HMI tags "VAT_DB_SDC_EMS_FLAGS"
   "SDC\DB_SDC_EMS_FLAGS\DB_SDC_EMS_FLAGS.EMS[8]" : Int AT %DB0.DBW0, 1 s   // EMSdriver present
   "SDC\DB_SDC_EMS_FLAGS\_EMS_Flags_HMI_Byte_00" : Int, internal
   "SDC\DB_SDC_EMS_FLAGS\_EMS_Flags_HMI_Byte_19" : Int, internal
   "DB_SDC_EMS_FLAGS_HMI_HMI[1].RET_VAL_SFC12" : Int = PLC DB_SDC_EMS_FLAGS_HMI.HMI[1].RET_VAL_SFC12 AT %DB3801.DBW34, 1 s   // RetVal SFC12
   "SDC\DB_SDC_EMS_FLAGS\DB_SDC_EMS_FLAGS.EMS[9]" : Int AT %DB0.DBW0, 1 s   // EMSdriver present
   "SDC\DB_SDC_EMS_FLAGS\DB_SDC_EMS_FLAGS.EMS[19]" : Int AT %DB0.DBW0, 1 s   // EMSdriver present
   "SDC\DB_SDC_EMS_FLAGS\DB_SDC_EMS_FLAGS.HMI[XX].EMS_Nr" : Int AT %DB0.DBW0, 1 s   // Sektionsnummer
   "SDC\DB_SDC_EMS_FLAGS\_EMS_Flags_HMI_Byte_04" : Int, internal
   "SDC\DB_SDC_EMS_FLAGS\DB_SDC_EMS_FLAGS.HMI[XX].PULT_Nr_EDIT" : Int AT %DB0.DBW0, 1 s   // Pult Nr Editieren Aktiv (HMI 1 = Master)
   "SDC\DB_SDC_EMS_FLAGS\DB_SDC_EMS_FLAGS.EMS[20]" : Int AT %DB0.DBW0, 1 s   // EMSdriver present
   "DB_SDC_EMS_FLAGS_HEADER.LAENGE_EMS_FLAGS" : Int = PLC DB_SDC_EMS_FLAGS.HEADER.LAENGE_EMS_FLAGS AT %DB3701.DBW8, 1 s   // Länge Eingänge pro EMS
   "SDC\DB_SDC_EMS_FLAGS\DB_SDC_EMS_FLAGS.EMS[6]" : Int AT %DB0.DBW0, 1 s   // EMSdriver present
   "SDC\DB_SDC_EMS_FLAGS\DB_SDC_EMS_FLAGS.EMS[12]" : Int AT %DB0.DBW0, 1 s   // EMSdriver present
   "SDC\DB_SDC_EMS_FLAGS\DB_SDC_EMS_FLAGS.EMS[1]" : Int AT %DB0.DBW0, 1 s   // EMSdriver present
   "SDC\DB_SDC_EMS_FLAGS\DB_SDC_EMS_FLAGS.EMS[3]" : Int AT %DB0.DBW0, 1 s   // EMSdriver present
   "SDC\DB_SDC_EMS_FLAGS\DB_SDC_EMS_FLAGS.HMI[XX].BILD_Nr" : Int AT %DB0.DBW0, 1 s   // Bild_Nr aktiv
   "SDC\DB_SDC_EMS_FLAGS\DB_SDC_EMS_FLAGS.HMI[XX].T_LOAD" : Bool AT %DB0.DBX0.3, 1 s   // Taster laden
   "DB_SDC_EMS_FLAGS_HMI_HEADER.START_HMI" : Int = PLC DB_SDC_EMS_FLAGS_HMI.HEADER.START_HMI AT %DB3801.DBW10, 1 s   // Startadresse HMI
   "SDC\DB_SDC_EMS_FLAGS\DB_SDC_EMS_FLAGS.EMS[10]" : Int AT %DB0.DBW0, 1 s   // EMSdriver present
   "SDC\DB_SDC_EMS_FLAGS\_EMS_Flags_HMI_Byte_18" : Int, internal
   "SDC\DB_SDC_EMS_FLAGS\DB_SDC_EMS_FLAGS.EMS[7]" : Int AT %DB0.DBW0, 1 s   // EMSdriver present
   "SDC\DB_SDC_EMS_FLAGS\DB_SDC_EMS_FLAGS.EMS[13]" : Int AT %DB0.DBW0, 1 s   // EMSdriver present
   "DB_SDC_EMS_FLAGS_HMI_HMI[1].MODE_SFC12" : Byte = PLC DB_SDC_EMS_FLAGS_HMI.HMI[1].MODE_SFC12 AT %DB3801.DBB36, 1 s   // Mode SFC12
   "SDC\DB_SDC_EMS_FLAGS\DB_SDC_EMS_FLAGS.HMI[XX].FR_EDIT" : Bool AT %DB0.DBX0.0, 1 s   // Freigabe Editieren
   "SDC\DB_SDC_EMS_FLAGS\_EMS_Flags_HMI_Byte_12" : Int, internal
   "SDC\DB_SDC_EMS_FLAGS\DB_SDC_EMS_FLAGS.EMS[18]" : Int AT %DB0.DBW0, 1 s   // EMSdriver present
   "DB_SDC_EMS_FLAGS_HEADER.DB_NR" : Int = PLC DB_SDC_EMS_FLAGS.HEADER.DB_NR AT %DB3701.DBW0, 1 s   // DB Nummer
   "SDC\DB_SDC_EMS_FLAGS\DB_SDC_EMS_FLAGS.HMI[XX].BILD_Nr_Alt" : Int AT %DB0.DBW0, 1 s   // Bild_Nr alt
   "DB_SDC_EMS_FLAGS_HMI_HEADER.OFFEST_HMI_DATA" : Int = PLC DB_SDC_EMS_FLAGS_HMI.HEADER.OFFEST_HMI_DATA AT %DB3801.DBW12, 1 s   // Offestadresse der HMI Flag Data
   "SDC\DB_SDC_EMS_FLAGS\DB_SDC_EMS_FLAGS.EMS[2]" : Int AT %DB0.DBW0, 1 s   // EMSdriver present
   "DB_SDC_EMS_FLAGS_HEADER.MIN_NR_EMS" : Int = PLC DB_SDC_EMS_FLAGS.HEADER.MIN_NR_EMS AT %DB3701.DBW2, 1 s   // Niedrigste EMS Nummer im Daten DB
   "SDC\DB_SDC_EMS_FLAGS\DB_SDC_EMS_FLAGS.HMI[XX].T_ACTIV" : Bool AT %DB0.DBX0.4, 1 s   // Taster activieren
   "SDC\DB_SDC_EMS_FLAGS\DB_SDC_EMS_FLAGS.EMS[16]" : Int AT %DB0.DBW0, 1 s   // EMSdriver present
   "SDC\DB_SDC_EMS_FLAGS\DB_SDC_EMS_FLAGS.HMI[XX].T_DEACTIV" : Bool AT %DB0.DBX0.5, 1 s   // Taster deactivieren
   "DB_SDC_EMS_FLAGS_HEADER.MAX_NR_EMS" : Int = PLC DB_SDC_EMS_FLAGS.HEADER.MAX_NR_EMS AT %DB3701.DBW4, 1 s   // Höchste EMS Nummer im Daten DB
   "DB_SDC_EMS_FLAGS_HMI_HMI[1].REQ_SFC12" : Bool = PLC DB_SDC_EMS_FLAGS_HMI.HMI[1].REQ_SFC12 AT %DB3801.DBX39.3, 1 s   // Request SFC12
   "SDC\DB_SDC_EMS_FLAGS\DB_SDC_EMS_FLAGS.HMI[XX].T_RESET_BED" : Bool AT %DB0.DBX0.1, 1 s   // Taster Reset Bedienfreigabe Pult Nr Bedienung
   "SDC\DB_SDC_EMS_FLAGS\_EMS_Flags_HMI_Byte_20" : Int, internal
   "DB_SDC_EMS_FLAGS_HMI_HMI[1].PULT_Nr_EDIT" : Int = PLC DB_SDC_EMS_FLAGS_HMI.HMI[1].PULT_Nr_EDIT AT %DB3801.DBW20, 1 s   // Pult Nr Editieren Aktiv (HMI 1 = Master)
   "SDC\DB_SDC_EMS_FLAGS\DB_SDC_EMS_FLAGS.HMI[XX].ER_DATA" : Bool AT %DB0.DBX0.1, 1 s   // Daten Fehlerhaft
   "SDC\DB_SDC_EMS_FLAGS\_EMS_Flags_HMI_Byte_08" : Int, internal
   "SDC\DB_SDC_EMS_FLAGS\DB_SDC_EMS_FLAGS.EMS[11]" : Int AT %DB0.DBW0, 1 s   // EMSdriver present
   "DB_SDC_EMS_FLAGS_HMI_HMI[1].TIME_SFC12" : Int = PLC DB_SDC_EMS_FLAGS_HMI.HMI[1].TIME_SFC12 AT %DB3801.DBW30, 1 s   // Actuelle Zeit Activieren/Deactivieren
   "SDC\DB_SDC_EMS_FLAGS\DB_SDC_EMS_FLAGS.EMS[14]" : Int AT %DB0.DBW0, 1 s   // EMSdriver present
   "SDC\DB_SDC_EMS_FLAGS\_EMS_Flags_HMI_Byte_16" : Int, internal
   "SDC\DB_SDC_EMS_FLAGS\DB_SDC_EMS_FLAGS.HMI[XX].T_SAVE" : Bool AT %DB0.DBX0.2, 1 s   // Taster speichern
   "SDC\DB_SDC_EMS_FLAGS\DB_SDC_EMS_FLAGS.EMS[15]" : Int AT %DB0.DBW0, 1 s   // EMSdriver present
   "SDC\DB_SDC_EMS_FLAGS\_EMS_Flags_HMI_Byte_10" : Int, internal
   "SDC\DB_SDC_EMS_FLAGS\_EMS_Flags_HMI_Byte_14" : Int, internal
   "SDC\DB_SDC_EMS_FLAGS\DB_SDC_EMS_FLAGS.HMI[XX].T_EDIT" : Bool AT %DB0.DBX0.0, 1 s   // Taster Editieren für Pult aktivieren
   "SDC\DB_SDC_EMS_FLAGS\_EMS_Flags_HMI_Byte_09" : Int, internal
   "DB_SDC_EMS_FLAGS_HMI_HMI[1].BUSY_SFC12" : Bool = PLC DB_SDC_EMS_FLAGS_HMI.HMI[1].BUSY_SFC12 AT %DB3801.DBX39.2, 1 s   // Busy SFC12
   "SDC\DB_SDC_EMS_FLAGS\_EMS_Nr" : Int, internal
      on ChangeValue: "SDC_TS_PARAMETER"(); "SDC_TS_REFERENCE"("SDC\DB_SDC_EMS_FLAGS\_EMS_Nr")
   "SDC\DB_SDC_EMS_FLAGS\DB_SDC_EMS_FLAGS.EMS[17]" : Int AT %DB0.DBW0, 1 s   // EMSdriver present
   "SDC\DB_SDC_EMS_FLAGS\_EMS_Flags_HMI_Byte_06" : Int, internal
   "SDC\DB_SDC_EMS_FLAGS\DB_SDC_EMS_FLAGS.HMI[XX].FLAGS" : Word AT %DB0.DBW0, 1 s   // Freigabe Editieren
   "SDC\DB_SDC_EMS_FLAGS\_EMS_Flags_HMI_Byte_02" : Int, internal
   "SDC\DB_SDC_EMS_FLAGS\DB_SDC_EMS_FLAGS.EMS[5]" : Int AT %DB0.DBW0, 1 s   // EMSdriver present
   "DB_SDC_EMS_FLAGS_HEADER.START_EMS" : Int = PLC DB_SDC_EMS_FLAGS.HEADER.START_EMS AT %DB3701.DBW6, 1 s   // Startadresse der EMS Daten im Daten DB
   "SDC\DB_SDC_EMS_FLAGS\DB_SDC_EMS_FLAGS.EMS[4]" : Int AT %DB0.DBW0, 1 s   // EMSdriver present
   "SDC\DB_SDC_EMS_FLAGS\DB_SDC_EMS_FLAGS.HMI[1].LADDR_SFC12" : Int AT %DB0.DBW32, 1 s   // Actuelle LADDR
   "SDC\DB_SDC_EMS_FLAGS\DB_SDC_EMS_FLAGS.EMS[21]" : Int AT %DB0.DBW0, 1 s   // EMSdriver present
   "SDC\DB_SDC_EMS_FLAGS\DB_SDC_EMS_FLAGS.EMS[22]" : Int AT %DB0.DBW0, 1 s
   "SDC\DB_SDC_EMS_FLAGS\DB_SDC_EMS_FLAGS.EMS[23]" : Int AT %DB0.DBW0, 1 s
   "SDC\DB_SDC_EMS_FLAGS\DB_SDC_EMS_FLAGS.EMS[24]" : Int AT %DB0.DBW0, 1 s
   "SDC\DB_SDC_EMS_FLAGS\DB_SDC_EMS_FLAGS.EMS[25]" : Int AT %DB0.DBW0, 1 s
   "SDC\DB_SDC_EMS_FLAGS\DB_SDC_EMS_FLAGS.EMS[26]" : Int AT %DB0.DBW0, 1 s
   "SDC\DB_SDC_EMS_FLAGS\DB_SDC_EMS_FLAGS.EMS[27]" : Int AT %DB0.DBW0, 1 s
   "SDC\DB_SDC_EMS_FLAGS\DB_SDC_EMS_FLAGS.EMS[28]" : Int AT %DB0.DBW0, 1 s
   "SDC\DB_SDC_EMS_FLAGS\DB_SDC_EMS_FLAGS.EMS[29]" : Int AT %DB0.DBW0, 1 s
   "SDC\DB_SDC_EMS_FLAGS\DB_SDC_EMS_FLAGS.EMS[30]" : Int AT %DB0.DBW0, 1 s
   "SDC\DB_SDC_EMS_FLAGS\DB_SDC_EMS_FLAGS.EMS[31]" : Int AT %DB0.DBW0, 1 s
   "SDC\DB_SDC_EMS_FLAGS\DB_SDC_EMS_FLAGS.EMS[32]" : Int AT %DB0.DBW0, 1 s
   "SDC\DB_SDC_EMS_FLAGS\DB_SDC_EMS_FLAGS.EMS[33]" : Int AT %DB0.DBW0, 1 s
   "SDC\DB_SDC_EMS_FLAGS\DB_SDC_EMS_FLAGS.EMS[34]" : Int AT %DB0.DBW0, 1 s
   "SDC\DB_SDC_EMS_FLAGS\DB_SDC_EMS_FLAGS.EMS[35]" : Int AT %DB0.DBW0, 1 s
   "SDC\DB_SDC_EMS_FLAGS\DB_SDC_EMS_FLAGS.EMS[36]" : Int AT %DB0.DBW0, 1 s
   "SDC\DB_SDC_EMS_FLAGS\DB_SDC_EMS_FLAGS.EMS[37]" : Int AT %DB0.DBW0, 1 s
   "SDC\DB_SDC_EMS_FLAGS\DB_SDC_EMS_FLAGS.EMS[38]" : Int AT %DB0.DBW0, 1 s
   "SDC\DB_SDC_EMS_FLAGS\DB_SDC_EMS_FLAGS.EMS[39]" : Int AT %DB0.DBW0, 1 s
   "SDC\DB_SDC_EMS_FLAGS\DB_SDC_EMS_FLAGS.EMS[40]" : Int AT %DB0.DBW0, 1 s
   "SDC\DB_SDC_EMS_FLAGS\DB_SDC_EMS_FLAGS.EMS[41]" : Int AT %DB0.DBW0, 1 s
   "SDC\DB_SDC_EMS_FLAGS\DB_SDC_EMS_FLAGS.EMS[42]" : Int AT %DB0.DBW0, 1 s
   "SDC\DB_SDC_EMS_FLAGS\DB_SDC_EMS_FLAGS.EMS[43]" : Int AT %DB0.DBW0, 1 s
   "SDC\DB_SDC_EMS_FLAGS\DB_SDC_EMS_FLAGS.EMS[44]" : Int AT %DB0.DBW0, 1 s
   "SDC\DB_SDC_EMS_FLAGS\DB_SDC_EMS_FLAGS.EMS[45]" : Int AT %DB0.DBW0, 1 s
   "SDC\DB_SDC_EMS_FLAGS\DB_SDC_EMS_FLAGS.EMS[46]" : Int AT %DB0.DBW0, 1 s
   "SDC\DB_SDC_EMS_FLAGS\DB_SDC_EMS_FLAGS.EMS[47]" : Int AT %DB0.DBW0, 1 s
   "SDC\DB_SDC_EMS_FLAGS\DB_SDC_EMS_FLAGS.EMS[48]" : Int AT %DB0.DBW0, 1 s
   "SDC\DB_SDC_EMS_FLAGS\DB_SDC_EMS_FLAGS.EMS[49]" : Int AT %DB0.DBW0, 1 s
   "SDC\DB_SDC_EMS_FLAGS\DB_SDC_EMS_FLAGS.EMS[50]" : Int AT %DB0.DBW0, 1 s
   "SDC\DB_SDC_EMS_FLAGS\DB_SDC_EMS_FLAGS.EMS[51]" : Int AT %DB0.DBW0, 1 s
   "SDC\DB_SDC_EMS_FLAGS\DB_SDC_EMS_FLAGS.EMS[52]" : Int AT %DB0.DBW0, 1 s
   "SDC\DB_SDC_EMS_FLAGS\DB_SDC_EMS_FLAGS.EMS[53]" : Int AT %DB0.DBW0, 1 s
   "SDC\DB_SDC_EMS_FLAGS\DB_SDC_EMS_FLAGS.EMS[54]" : Int AT %DB0.DBW0, 1 s
   "SDC\DB_SDC_EMS_FLAGS\DB_SDC_EMS_FLAGS.EMS[55]" : Int AT %DB0.DBW0, 1 s
   "SDC\DB_SDC_EMS_FLAGS\DB_SDC_EMS_FLAGS.EMS[56]" : Int AT %DB0.DBW0, 1 s
   "SDC\DB_SDC_EMS_FLAGS\DB_SDC_EMS_FLAGS.EMS[57]" : Int AT %DB0.DBW0, 1 s
   "SDC\DB_SDC_EMS_FLAGS\DB_SDC_EMS_FLAGS.EMS[58]" : Int AT %DB0.DBW0, 1 s
   "SDC\DB_SDC_EMS_FLAGS\DB_SDC_EMS_FLAGS.EMS[59]" : Int AT %DB0.DBW0, 1 s
   "SDC\DB_SDC_EMS_FLAGS\DB_SDC_EMS_FLAGS.EMS[60]" : Int AT %DB0.DBW0, 1 s
   "SDC\DB_SDC_EMS_FLAGS\DB_SDC_EMS_FLAGS.EMS[61]" : Int AT %DB0.DBW0, 1 s
   "SDC\DB_SDC_EMS_FLAGS\DB_SDC_EMS_FLAGS.EMS[62]" : Int AT %DB0.DBW0, 1 s
   "SDC\DB_SDC_EMS_FLAGS\DB_SDC_EMS_FLAGS.EMS[63]" : Int AT %DB0.DBW0, 1 s
   "SDC\DB_SDC_EMS_FLAGS\DB_SDC_EMS_FLAGS.EMS[64]" : Int AT %DB0.DBW0, 1 s
   "SDC\DB_SDC_EMS_FLAGS\DB_SDC_EMS_FLAGS.EMS[65]" : Int AT %DB0.DBW0, 1 s
   "SDC\DB_SDC_EMS_FLAGS\DB_SDC_EMS_FLAGS.EMS[66]" : Int AT %DB0.DBW0, 1 s
   "SDC\DB_SDC_EMS_FLAGS\DB_SDC_EMS_FLAGS.EMS[67]" : Int AT %DB0.DBW0, 1 s
   "SDC\DB_SDC_EMS_FLAGS\DB_SDC_EMS_FLAGS.EMS[68]" : Int AT %DB0.DBW0, 1 s
   "SDC\DB_SDC_EMS_FLAGS\DB_SDC_EMS_FLAGS.EMS[69]" : Int AT %DB0.DBW0, 1 s
   "SDC\DB_SDC_EMS_FLAGS\DB_SDC_EMS_FLAGS.EMS[70]" : Int AT %DB0.DBW0, 1 s
   "SDC\DB_SDC_EMS_FLAGS\DB_SDC_EMS_FLAGS.EMS[71]" : Int AT %DB0.DBW0, 1 s
   "SDC\DB_SDC_EMS_FLAGS\DB_SDC_EMS_FLAGS.EMS[72]" : Int AT %DB0.DBW0, 1 s
   "SDC\DB_SDC_EMS_FLAGS\DB_SDC_EMS_FLAGS.EMS[73]" : Int AT %DB0.DBW0, 1 s
   "SDC\DB_SDC_EMS_FLAGS\DB_SDC_EMS_FLAGS.EMS[74]" : Int AT %DB0.DBW0, 1 s
   "SDC\DB_SDC_EMS_FLAGS\DB_SDC_EMS_FLAGS.EMS[75]" : Int AT %DB0.DBW0, 1 s
   "SDC\DB_SDC_EMS_FLAGS\DB_SDC_EMS_FLAGS.EMS[76]" : Int AT %DB0.DBW0, 1 s
   "SDC\DB_SDC_EMS_FLAGS\DB_SDC_EMS_FLAGS.EMS[77]" : Int AT %DB0.DBW0, 1 s
   "SDC\DB_SDC_EMS_FLAGS\DB_SDC_EMS_FLAGS.EMS[78]" : Int AT %DB0.DBW0, 1 s
   "SDC\DB_SDC_EMS_FLAGS\DB_SDC_EMS_FLAGS.EMS[79]" : Int AT %DB0.DBW0, 1 s
   "SDC\DB_SDC_EMS_FLAGS\DB_SDC_EMS_FLAGS.EMS[80]" : Int AT %DB0.DBW0, 1 s
   "SDC\DB_SDC_EMS_FLAGS\DB_SDC_EMS_FLAGS.EMS[81]" : Int AT %DB0.DBW0, 1 s
   "SDC\DB_SDC_EMS_FLAGS\DB_SDC_EMS_FLAGS.EMS[82]" : Int AT %DB0.DBW0, 1 s
   "SDC\DB_SDC_EMS_FLAGS\DB_SDC_EMS_FLAGS.EMS[83]" : Int AT %DB0.DBW0, 1 s
   "SDC\DB_SDC_EMS_FLAGS\DB_SDC_EMS_FLAGS.EMS[84]" : Int AT %DB0.DBW0, 1 s
   "SDC\DB_SDC_EMS_FLAGS\DB_SDC_EMS_FLAGS.EMS[85]" : Int AT %DB0.DBW0, 1 s
   "SDC\DB_SDC_EMS_FLAGS\DB_SDC_EMS_FLAGS.EMS[86]" : Int AT %DB0.DBW0, 1 s
   "SDC\DB_SDC_EMS_FLAGS\DB_SDC_EMS_FLAGS.EMS[87]" : Int AT %DB0.DBW0, 1 s
   "SDC\DB_SDC_EMS_FLAGS\DB_SDC_EMS_FLAGS.EMS[88]" : Int AT %DB0.DBW0, 1 s
   "SDC\DB_SDC_EMS_FLAGS\DB_SDC_EMS_FLAGS.EMS[89]" : Int AT %DB0.DBW0, 1 s
   "SDC\DB_SDC_EMS_FLAGS\DB_SDC_EMS_FLAGS.EMS[90]" : Int AT %DB0.DBW0, 1 s
   "SDC\DB_SDC_EMS_FLAGS\DB_SDC_EMS_FLAGS.EMS[91]" : Int AT %DB0.DBW0, 1 s
   "SDC\DB_SDC_EMS_FLAGS\DB_SDC_EMS_FLAGS.EMS[92]" : Int AT %DB0.DBW0, 1 s
   "SDC\DB_SDC_EMS_FLAGS\DB_SDC_EMS_FLAGS.EMS[93]" : Int AT %DB0.DBW0, 1 s
   "SDC\DB_SDC_EMS_FLAGS\DB_SDC_EMS_FLAGS.EMS[94]" : Int AT %DB0.DBW0, 1 s
   "SDC\DB_SDC_EMS_FLAGS\DB_SDC_EMS_FLAGS.EMS[95]" : Int AT %DB0.DBW0, 1 s
   "SDC\DB_SDC_EMS_FLAGS\DB_SDC_EMS_FLAGS.EMS[96]" : Int AT %DB0.DBW0, 1 s
   "SDC\DB_SDC_EMS_FLAGS\DB_SDC_EMS_FLAGS.EMS[97]" : Int AT %DB0.DBW0, 1 s
   "SDC\DB_SDC_EMS_FLAGS\DB_SDC_EMS_FLAGS.EMS[98]" : Int AT %DB0.DBW0, 1 s
   "SDC\DB_SDC_EMS_FLAGS\DB_SDC_EMS_FLAGS.EMS[99]" : Int AT %DB0.DBW0, 1 s
   "SDC\DB_SDC_EMS_FLAGS\DB_SDC_EMS_FLAGS.EMS[100]" : Int AT %DB0.DBW0, 1 s
   "SDC\DB_SDC_EMS_FLAGS\DB_SDC_EMS_FLAGS.EMS[101]" : Int AT %DB0.DBW0, 1 s
   "SDC\DB_SDC_EMS_FLAGS\DB_SDC_EMS_FLAGS.EMS[102]" : Int AT %DB0.DBW0, 1 s
   "SDC\DB_SDC_EMS_FLAGS\DB_SDC_EMS_FLAGS.EMS[103]" : Int AT %DB0.DBW0, 1 s
   "SDC\DB_SDC_EMS_FLAGS\DB_SDC_EMS_FLAGS.EMS[104]" : Int AT %DB0.DBW0, 1 s
   "SDC\DB_SDC_EMS_FLAGS\DB_SDC_EMS_FLAGS.EMS[105]" : Int AT %DB0.DBW0, 1 s
   "SDC\DB_SDC_EMS_FLAGS\DB_SDC_EMS_FLAGS.EMS[106]" : Int AT %DB0.DBW0, 1 s
   "SDC\DB_SDC_EMS_FLAGS\DB_SDC_EMS_FLAGS.EMS[107]" : Int AT %DB0.DBW0, 1 s
   "SDC\DB_SDC_EMS_FLAGS\DB_SDC_EMS_FLAGS.EMS[108]" : Int AT %DB0.DBW0, 1 s
   "SDC\DB_SDC_EMS_FLAGS\DB_SDC_EMS_FLAGS.EMS[109]" : Int AT %DB0.DBW0, 1 s
   "SDC\DB_SDC_EMS_FLAGS\_EMS_Flags_Byte_EMS001" : Int, internal
   "SDC\DB_SDC_EMS_FLAGS\_EMS_Flags_Byte_EMS002" : Int, internal
   "SDC\DB_SDC_EMS_FLAGS\_EMS_Flags_Byte_EMS003" : Int, internal
   "SDC\DB_SDC_EMS_FLAGS\_EMS_Flags_Byte_EMS004" : Int, internal
   "SDC\DB_SDC_EMS_FLAGS\_EMS_Flags_Byte_EMS005" : Int, internal
   "SDC\DB_SDC_EMS_FLAGS\_EMS_Flags_Byte_EMS006" : Int, internal
   "SDC\DB_SDC_EMS_FLAGS\_EMS_Flags_Byte_EMS007" : Int, internal
   "SDC\DB_SDC_EMS_FLAGS\_EMS_Flags_Byte_EMS008" : Int, internal
   "SDC\DB_SDC_EMS_FLAGS\_EMS_Flags_Byte_EMS009" : Int, internal
   "SDC\DB_SDC_EMS_FLAGS\_EMS_Flags_Byte_EMS010" : Int, internal
   "SDC\DB_SDC_EMS_FLAGS\_EMS_Flags_Byte_EMS011" : Int, internal
   "SDC\DB_SDC_EMS_FLAGS\_EMS_Flags_Byte_EMS012" : Int, internal
   "SDC\DB_SDC_EMS_FLAGS\_EMS_Flags_Byte_EMS013" : Int, internal
   "SDC\DB_SDC_EMS_FLAGS\_EMS_Flags_Byte_EMS014" : Int, internal
   "SDC\DB_SDC_EMS_FLAGS\_EMS_Flags_Byte_EMS015" : Int, internal
   "SDC\DB_SDC_EMS_FLAGS\_EMS_Flags_Byte_EMS016" : Int, internal
   "SDC\DB_SDC_EMS_FLAGS\_EMS_Flags_Byte_EMS017" : Int, internal
   "SDC\DB_SDC_EMS_FLAGS\_EMS_Flags_Byte_EMS018" : Int, internal
   "SDC\DB_SDC_EMS_FLAGS\_EMS_Flags_Byte_EMS019" : Int, internal
   "SDC\DB_SDC_EMS_FLAGS\_EMS_Flags_Byte_EMS020" : Int, internal
   "SDC\DB_SDC_EMS_FLAGS\_EMS_Flags_Byte_EMS021" : Int, internal
   "SDC\DB_SDC_EMS_FLAGS\_EMS_Flags_Byte_EMS022" : Int, internal
   "SDC\DB_SDC_EMS_FLAGS\_EMS_Flags_Byte_EMS023" : Int, internal
   "SDC\DB_SDC_EMS_FLAGS\_EMS_Flags_Byte_EMS024" : Int, internal
   "SDC\DB_SDC_EMS_FLAGS\_EMS_Flags_Byte_EMS025" : Int, internal
   "SDC\DB_SDC_EMS_FLAGS\_EMS_Flags_Byte_EMS026" : Int, internal
   "SDC\DB_SDC_EMS_FLAGS\_EMS_Flags_Byte_EMS027" : Int, internal
   "SDC\DB_SDC_EMS_FLAGS\_EMS_Flags_Byte_EMS028" : Int, internal
   "SDC\DB_SDC_EMS_FLAGS\_EMS_Flags_Byte_EMS029" : Int, internal
   "SDC\DB_SDC_EMS_FLAGS\_EMS_Flags_Byte_EMS030" : Int, internal
   "SDC\DB_SDC_EMS_FLAGS\_EMS_Flags_Byte_EMS031" : Int, internal
   "SDC\DB_SDC_EMS_FLAGS\_EMS_Flags_Byte_EMS032" : Int, internal
   "SDC\DB_SDC_EMS_FLAGS\_EMS_Flags_Byte_EMS033" : Int, internal
   "SDC\DB_SDC_EMS_FLAGS\_EMS_Flags_Byte_EMS034" : Int, internal
   "SDC\DB_SDC_EMS_FLAGS\_EMS_Flags_Byte_EMS035" : Int, internal
   "SDC\DB_SDC_EMS_FLAGS\_EMS_Flags_Byte_EMS036" : Int, internal
   "SDC\DB_SDC_EMS_FLAGS\_EMS_Flags_Byte_EMS037" : Int, internal
   "SDC\DB_SDC_EMS_FLAGS\_EMS_Flags_Byte_EMS038" : Int, internal
   "SDC\DB_SDC_EMS_FLAGS\_EMS_Flags_Byte_EMS039" : Int, internal
   "SDC\DB_SDC_EMS_FLAGS\_EMS_Flags_Byte_EMS040" : Int, internal
   "SDC\DB_SDC_EMS_FLAGS\_EMS_Flags_Byte_EMS041" : Int, internal
   "SDC\DB_SDC_EMS_FLAGS\_EMS_Flags_Byte_EMS042" : Int, internal
   "SDC\DB_SDC_EMS_FLAGS\_EMS_Flags_Byte_EMS043" : Int, internal
   "SDC\DB_SDC_EMS_FLAGS\_EMS_Flags_Byte_EMS044" : Int, internal
   "SDC\DB_SDC_EMS_FLAGS\_EMS_Flags_Byte_EMS045" : Int, internal
   "SDC\DB_SDC_EMS_FLAGS\_EMS_Flags_Byte_EMS046" : Int, internal
   "SDC\DB_SDC_EMS_FLAGS\_EMS_Flags_Byte_EMS047" : Int, internal
   "SDC\DB_SDC_EMS_FLAGS\_EMS_Flags_Byte_EMS048" : Int, internal
   "SDC\DB_SDC_EMS_FLAGS\_EMS_Flags_Byte_EMS049" : Int, internal
   "SDC\DB_SDC_EMS_FLAGS\_EMS_Flags_Byte_EMS050" : Int, internal
   "SDC\DB_SDC_EMS_FLAGS\_EMS_Flags_Byte_EMS051" : Int, internal
   "SDC\DB_SDC_EMS_FLAGS\_EMS_Flags_Byte_EMS052" : Int, internal
   "SDC\DB_SDC_EMS_FLAGS\_EMS_Flags_Byte_EMS053" : Int, internal
   "SDC\DB_SDC_EMS_FLAGS\_EMS_Flags_Byte_EMS054" : Int, internal
   "SDC\DB_SDC_EMS_FLAGS\_EMS_Flags_Byte_EMS055" : Int, internal
   "SDC\DB_SDC_EMS_FLAGS\_EMS_Flags_Byte_EMS056" : Int, internal
   "SDC\DB_SDC_EMS_FLAGS\_EMS_Flags_Byte_EMS057" : Int, internal
   "SDC\DB_SDC_EMS_FLAGS\_EMS_Flags_Byte_EMS058" : Int, internal
   "SDC\DB_SDC_EMS_FLAGS\_EMS_Flags_Byte_EMS059" : Int, internal
   "SDC\DB_SDC_EMS_FLAGS\_EMS_Flags_Byte_EMS060" : Int, internal
   "SDC\DB_SDC_EMS_FLAGS\_EMS_Flags_Byte_EMS061" : Int, internal
   "SDC\DB_SDC_EMS_FLAGS\_EMS_Flags_Byte_EMS062" : Int, internal
   "SDC\DB_SDC_EMS_FLAGS\_EMS_Flags_Byte_EMS063" : Int, internal
   "SDC\DB_SDC_EMS_FLAGS\_EMS_Flags_Byte_EMS064" : Int, internal
   "SDC\DB_SDC_EMS_FLAGS\_EMS_Flags_Byte_EMS065" : Int, internal
   "SDC\DB_SDC_EMS_FLAGS\_EMS_Flags_Byte_EMS066" : Int, internal
   "SDC\DB_SDC_EMS_FLAGS\_EMS_Flags_Byte_EMS067" : Int, internal
   "SDC\DB_SDC_EMS_FLAGS\_EMS_Flags_Byte_EMS068" : Int, internal
   "SDC\DB_SDC_EMS_FLAGS\_EMS_Flags_Byte_EMS069" : Int, internal
   "SDC\DB_SDC_EMS_FLAGS\_EMS_Flags_Byte_EMS070" : Int, internal
   "SDC\DB_SDC_EMS_FLAGS\_EMS_Flags_Byte_EMS071" : Int, internal
   "SDC\DB_SDC_EMS_FLAGS\_EMS_Flags_Byte_EMS072" : Int, internal
   "SDC\DB_SDC_EMS_FLAGS\_EMS_Flags_Byte_EMS073" : Int, internal
   "SDC\DB_SDC_EMS_FLAGS\_EMS_Flags_Byte_EMS074" : Int, internal
   "SDC\DB_SDC_EMS_FLAGS\_EMS_Flags_Byte_EMS075" : Int, internal
   "SDC\DB_SDC_EMS_FLAGS\_EMS_Flags_Byte_EMS076" : Int, internal
   "SDC\DB_SDC_EMS_FLAGS\_EMS_Flags_Byte_EMS077" : Int, internal
   "SDC\DB_SDC_EMS_FLAGS\_EMS_Flags_Byte_EMS078" : Int, internal
   "SDC\DB_SDC_EMS_FLAGS\_EMS_Flags_Byte_EMS079" : Int, internal
   "SDC\DB_SDC_EMS_FLAGS\_EMS_Flags_Byte_EMS080" : Int, internal
   "SDC\DB_SDC_EMS_FLAGS\_EMS_Flags_Byte_EMS081" : Int, internal
   "SDC\DB_SDC_EMS_FLAGS\_EMS_Flags_Byte_EMS082" : Int, internal
   "SDC\DB_SDC_EMS_FLAGS\_EMS_Flags_Byte_EMS083" : Int, internal
   "SDC\DB_SDC_EMS_FLAGS\_EMS_Flags_Byte_EMS084" : Int, internal
   "SDC\DB_SDC_EMS_FLAGS\_EMS_Flags_Byte_EMS085" : Int, internal
   "SDC\DB_SDC_EMS_FLAGS\_EMS_Flags_Byte_EMS086" : Int, internal
   "SDC\DB_SDC_EMS_FLAGS\_EMS_Flags_Byte_EMS087" : Int, internal
   "SDC\DB_SDC_EMS_FLAGS\_EMS_Flags_Byte_EMS088" : Int, internal
   "SDC\DB_SDC_EMS_FLAGS\_EMS_Flags_Byte_EMS089" : Int, internal
   "SDC\DB_SDC_EMS_FLAGS\_EMS_Flags_Byte_EMS090" : Int, internal
   "SDC\DB_SDC_EMS_FLAGS\_EMS_Flags_Byte_EMS091" : Int, internal
   "SDC\DB_SDC_EMS_FLAGS\_EMS_Flags_Byte_EMS092" : Int, internal
   "SDC\DB_SDC_EMS_FLAGS\_EMS_Flags_Byte_EMS093" : Int, internal
   "SDC\DB_SDC_EMS_FLAGS\_EMS_Flags_Byte_EMS094" : Int, internal
   "SDC\DB_SDC_EMS_FLAGS\_EMS_Flags_Byte_EMS095" : Int, internal
   "SDC\DB_SDC_EMS_FLAGS\_EMS_Flags_Byte_EMS096" : Int, internal
   "SDC\DB_SDC_EMS_FLAGS\_EMS_Flags_Byte_EMS097" : Int, internal
   "SDC\DB_SDC_EMS_FLAGS\_EMS_Flags_Byte_EMS098" : Int, internal
   "SDC\DB_SDC_EMS_FLAGS\_EMS_Flags_Byte_EMS099" : Int, internal
   "SDC\DB_SDC_EMS_FLAGS\_EMS_Flags_Byte_EMS100" : Int, internal
   "SDC\DB_SDC_EMS_FLAGS\_EMS_Flags_Byte_EMS101" : Int, internal
   "SDC\DB_SDC_EMS_FLAGS\_EMS_Flags_Byte_EMS102" : Int, internal
   "SDC\DB_SDC_EMS_FLAGS\_EMS_Flags_Byte_EMS103" : Int, internal
   "SDC\DB_SDC_EMS_FLAGS\_EMS_Flags_Byte_EMS104" : Int, internal
   "SDC\DB_SDC_EMS_FLAGS\_EMS_Flags_Byte_EMS105" : Int, internal
   "SDC\DB_SDC_EMS_FLAGS\_EMS_Flags_Byte_EMS106" : Int, internal
   "SDC\DB_SDC_EMS_FLAGS\_EMS_Flags_Byte_EMS107" : Int, internal
   "SDC\DB_SDC_EMS_FLAGS\_EMS_Flags_Byte_EMS108" : Int, internal
   "SDC\DB_SDC_EMS_FLAGS\_EMS_Flags_Byte_EMS109" : Int, internal
   "DB_SDC_EMS_FLAGS_HMI_HEADER.DB_NR" : Int = PLC DB_SDC_EMS_FLAGS_HMI.HEADER.DB_NR AT %DB3801.DBW0, 1 s
   "SDC\DB_SDC_EMS_FLAGS\_EMS_Flags_Byte_EMS110" : Int, internal
   "SDC\DB_SDC_EMS_FLAGS\_EMS_Flags_Byte_EMS111" : Int, internal
   "SDC\DB_SDC_EMS_FLAGS\_EMS_Flags_Byte_EMS112" : Int, internal
   "SDC\DB_SDC_EMS_FLAGS\_EMS_Flags_Byte_EMS113" : Int, internal
   "SDC\DB_SDC_EMS_FLAGS\_EMS_Flags_Byte_EMS114" : Int, internal
   "SDC\DB_SDC_EMS_FLAGS\_EMS_Flags_Byte_EMS115" : Int, internal
   "SDC\DB_SDC_EMS_FLAGS\_EMS_Flags_Byte_EMS116" : Int, internal
   "SDC\DB_SDC_EMS_FLAGS\_EMS_Flags_Byte_EMS117" : Int, internal
   "SDC\DB_SDC_EMS_FLAGS\_EMS_Flags_Byte_EMS118" : Int, internal
   "SDC\DB_SDC_EMS_FLAGS\_EMS_Flags_Byte_EMS119" : Int, internal
   "SDC\DB_SDC_EMS_FLAGS\_EMS_Flags_Byte_EMS120" : Int, internal
   "SDC\DB_SDC_EMS_FLAGS\_EMS_Flags_Byte_EMS121" : Int, internal
   "SDC\DB_SDC_EMS_FLAGS\_EMS_Flags_Byte_EMS122" : Int, internal
   "SDC\DB_SDC_EMS_FLAGS\_EMS_Flags_Byte_EMS123" : Int, internal
   "SDC\DB_SDC_EMS_FLAGS\_EMS_Flags_Byte_EMS124" : Int, internal
   "SDC\DB_SDC_EMS_FLAGS\_EMS_Flags_Byte_EMS125" : Int, internal
   "SDC\DB_SDC_EMS_FLAGS\_EMS_Flags_Byte_EMS126" : Int, internal
   "SDC\DB_SDC_EMS_FLAGS\_EMS_Flags_Byte_EMS127" : Int, internal
   "SDC\DB_SDC_EMS_FLAGS\_EMS_Flags_Byte_EMS128" : Int, internal
   "SDC\DB_SDC_EMS_FLAGS\_EMS_Flags_Byte_EMS129" : Int, internal
   "SDC\DB_SDC_EMS_FLAGS\_EMS_Flags_Byte_EMS130" : Int, internal
   "SDC\DB_SDC_EMS_FLAGS\_EMS_Flags_Byte_EMS131" : Int, internal
   "SDC\DB_SDC_EMS_FLAGS\_EMS_Flags_Byte_EMS132" : Int, internal
   "SDC\DB_SDC_EMS_FLAGS\_EMS_Flags_Byte_EMS133" : Int, internal
   "SDC\DB_SDC_EMS_FLAGS\_EMS_Flags_Byte_EMS134" : Int, internal
   "SDC\DB_SDC_EMS_FLAGS\_EMS_Flags_Byte_EMS135" : Int, internal
   "SDC\DB_SDC_EMS_FLAGS\_EMS_Flags_Byte_EMS136" : Int, internal
   "SDC\DB_SDC_EMS_FLAGS\_EMS_Flags_Byte_EMS137" : Int, internal
   "SDC\DB_SDC_EMS_FLAGS\_EMS_Flags_Byte_EMS138" : Int, internal
   "SDC\DB_SDC_EMS_FLAGS\_EMS_Flags_Byte_EMS139" : Int, internal
   "SDC\DB_SDC_EMS_FLAGS\_EMS_Flags_Byte_EMS140" : Int, internal
   "SDC\DB_SDC_EMS_FLAGS\_EMS_Flags_Byte_EMS141" : Int, internal
   "SDC\DB_SDC_EMS_FLAGS\_EMS_Flags_Byte_EMS142" : Int, internal
   "SDC\DB_SDC_EMS_FLAGS\_EMS_Flags_Byte_EMS143" : Int, internal
   "SDC\DB_SDC_EMS_FLAGS\_EMS_Flags_Byte_EMS144" : Int, internal
   "SDC\DB_SDC_EMS_FLAGS\_EMS_Flags_Byte_EMS145" : Int, internal
   "SDC\DB_SDC_EMS_FLAGS\_EMS_Flags_Byte_EMS146" : Int, internal
   "SDC\DB_SDC_EMS_FLAGS\_EMS_Flags_Byte_EMS147" : Int, internal
   "SDC\DB_SDC_EMS_FLAGS\_EMS_Flags_Byte_EMS148" : Int, internal
   "SDC\DB_SDC_EMS_FLAGS\_EMS_Flags_Byte_EMS149" : Int, internal
   "SDC\DB_SDC_EMS_FLAGS\_EMS_Flags_Byte_EMS150" : Int, internal
   "SDC\DB_SDC_EMS_FLAGS\_EMS_Flags_Byte_EMS151" : Int, internal
   "SDC\DB_SDC_EMS_FLAGS\_EMS_Flags_Byte_EMS152" : Int, internal
   "SDC\DB_SDC_EMS_FLAGS\_EMS_Flags_Byte_EMS153" : Int, internal
   "SDC\DB_SDC_EMS_FLAGS\_EMS_Flags_Byte_EMS154" : Int, internal
   "SDC\DB_SDC_EMS_FLAGS\_EMS_Flags_Byte_EMS155" : Int, internal
   "SDC\DB_SDC_EMS_FLAGS\_EMS_Flags_Byte_EMS156" : Int, internal
   "SDC\DB_SDC_EMS_FLAGS\_EMS_Flags_Byte_EMS157" : Int, internal
   "SDC\DB_SDC_EMS_FLAGS\_EMS_Flags_Byte_EMS158" : Int, internal
   "SDC\DB_SDC_EMS_FLAGS\_EMS_Flags_Byte_EMS159" : Int, internal
   "SDC\DB_SDC_EMS_FLAGS\_EMS_Flags_Byte_EMS160" : Int, internal
   "SDC\DB_SDC_EMS_FLAGS\_EMS_Flags_Byte_EMS161" : Int, internal
   "SDC\DB_SDC_EMS_FLAGS\_EMS_Flags_Byte_EMS162" : Int, internal
   "SDC\DB_SDC_EMS_FLAGS\_EMS_Flags_Byte_EMS163" : Int, internal
   "SDC\DB_SDC_EMS_FLAGS\_EMS_Flags_Byte_EMS164" : Int, internal
   "SDC\DB_SDC_EMS_FLAGS\_EMS_Flags_Byte_EMS165" : Int, internal
   "SDC\DB_SDC_EMS_FLAGS\_EMS_Flags_Byte_EMS166" : Int, internal
   "SDC\DB_SDC_EMS_FLAGS\_EMS_Flags_Byte_EMS167" : Int, internal
   "SDC\DB_SDC_EMS_FLAGS\_EMS_Flags_Byte_EMS168" : Int, internal
   "SDC\DB_SDC_EMS_FLAGS\_EMS_Flags_Byte_EMS169" : Int, internal
   "SDC\DB_SDC_EMS_FLAGS\_EMS_Flags_Byte_EMS170" : Int, internal
   "SDC\DB_SDC_EMS_FLAGS\_EMS_Flags_Byte_EMS171" : Int, internal
   "SDC\DB_SDC_EMS_FLAGS\_EMS_Flags_Byte_EMS172" : Int, internal
   "SDC\DB_SDC_EMS_FLAGS\_EMS_Flags_Byte_EMS173" : Int, internal
   "SDC\DB_SDC_EMS_FLAGS\_EMS_Flags_Byte_EMS174" : Int, internal
   "SDC\DB_SDC_EMS_FLAGS\_EMS_Flags_Byte_EMS175" : Int, internal
   "SDC\DB_SDC_EMS_FLAGS\_EMS_Flags_Byte_EMS176" : Int, internal
   "SDC\DB_SDC_EMS_FLAGS\_EMS_Flags_Byte_EMS177" : Int, internal
   "SDC\DB_SDC_EMS_FLAGS\_EMS_Flags_Byte_EMS178" : Int, internal
   "SDC\DB_SDC_EMS_FLAGS\_EMS_Flags_Byte_EMS179" : Int, internal
   "SDC\DB_SDC_EMS_FLAGS\_EMS_Flags_Byte_EMS180" : Int, internal
   "SDC\DB_SDC_EMS_FLAGS\_EMS_Flags_Byte_EMS181" : Int, internal
   "SDC\DB_SDC_EMS_FLAGS\_EMS_Flags_Byte_EMS182" : Int, internal
   "SDC\DB_SDC_EMS_FLAGS\_EMS_Flags_Byte_EMS183" : Int, internal
   "SDC\DB_SDC_EMS_FLAGS\_EMS_Flags_Byte_EMS184" : Int, internal
   "SDC\DB_SDC_EMS_FLAGS\DB_SDC_EMS_FLAGS.EMS[110]" : Int AT %DB0.DBW0, 1 s
   "SDC\DB_SDC_EMS_FLAGS\DB_SDC_EMS_FLAGS.EMS[111]" : Int AT %DB0.DBW0, 1 s
   "SDC\DB_SDC_EMS_FLAGS\DB_SDC_EMS_FLAGS.EMS[112]" : Int AT %DB0.DBW0, 1 s
   "SDC\DB_SDC_EMS_FLAGS\DB_SDC_EMS_FLAGS.EMS[113]" : Int AT %DB0.DBW0, 1 s
   "SDC\DB_SDC_EMS_FLAGS\DB_SDC_EMS_FLAGS.EMS[114]" : Int AT %DB0.DBW0, 1 s
   "SDC\DB_SDC_EMS_FLAGS\DB_SDC_EMS_FLAGS.EMS[115]" : Int AT %DB0.DBW0, 1 s
   "SDC\DB_SDC_EMS_FLAGS\DB_SDC_EMS_FLAGS.EMS[116]" : Int AT %DB0.DBW0, 1 s
   "SDC\DB_SDC_EMS_FLAGS\DB_SDC_EMS_FLAGS.EMS[117]" : Int AT %DB0.DBW0, 1 s
   "SDC\DB_SDC_EMS_FLAGS\DB_SDC_EMS_FLAGS.EMS[118]" : Int AT %DB0.DBW0, 1 s
   "SDC\DB_SDC_EMS_FLAGS\DB_SDC_EMS_FLAGS.EMS[119]" : Int AT %DB0.DBW0, 1 s
   "SDC\DB_SDC_EMS_FLAGS\DB_SDC_EMS_FLAGS.EMS[120]" : Int AT %DB0.DBW0, 1 s
   "SDC\DB_SDC_EMS_FLAGS\DB_SDC_EMS_FLAGS.EMS[121]" : Int AT %DB0.DBW0, 1 s
   "SDC\DB_SDC_EMS_FLAGS\DB_SDC_EMS_FLAGS.EMS[122]" : Int AT %DB0.DBW0, 1 s
   "SDC\DB_SDC_EMS_FLAGS\DB_SDC_EMS_FLAGS.EMS[123]" : Int AT %DB0.DBW0, 1 s
   "SDC\DB_SDC_EMS_FLAGS\DB_SDC_EMS_FLAGS.EMS[124]" : Int AT %DB0.DBW0, 1 s
   "SDC\DB_SDC_EMS_FLAGS\DB_SDC_EMS_FLAGS.EMS[125]" : Int AT %DB0.DBW0, 1 s
   "SDC\DB_SDC_EMS_FLAGS\DB_SDC_EMS_FLAGS.EMS[126]" : Int AT %DB0.DBW0, 1 s
   "SDC\DB_SDC_EMS_FLAGS\DB_SDC_EMS_FLAGS.EMS[127]" : Int AT %DB0.DBW0, 1 s
   "SDC\DB_SDC_EMS_FLAGS\DB_SDC_EMS_FLAGS.EMS[128]" : Int AT %DB0.DBW0, 1 s
   "SDC\DB_SDC_EMS_FLAGS\DB_SDC_EMS_FLAGS.EMS[129]" : Int AT %DB0.DBW0, 1 s
   "SDC\DB_SDC_EMS_FLAGS\DB_SDC_EMS_FLAGS.EMS[130]" : Int AT %DB0.DBW0, 1 s
   "SDC\DB_SDC_EMS_FLAGS\DB_SDC_EMS_FLAGS.EMS[131]" : Int AT %DB0.DBW0, 1 s
   "SDC\DB_SDC_EMS_FLAGS\DB_SDC_EMS_FLAGS.EMS[132]" : Int AT %DB0.DBW0, 1 s
   "SDC\DB_SDC_EMS_FLAGS\DB_SDC_EMS_FLAGS.EMS[133]" : Int AT %DB0.DBW0, 1 s
   "SDC\DB_SDC_EMS_FLAGS\DB_SDC_EMS_FLAGS.EMS[134]" : Int AT %DB0.DBW0, 1 s
   "SDC\DB_SDC_EMS_FLAGS\DB_SDC_EMS_FLAGS.EMS[135]" : Int AT %DB0.DBW0, 1 s
   "SDC\DB_SDC_EMS_FLAGS\DB_SDC_EMS_FLAGS.EMS[136]" : Int AT %DB0.DBW0, 1 s
   "SDC\DB_SDC_EMS_FLAGS\DB_SDC_EMS_FLAGS.EMS[137]" : Int AT %DB0.DBW0, 1 s
   "SDC\DB_SDC_EMS_FLAGS\DB_SDC_EMS_FLAGS.EMS[138]" : Int AT %DB0.DBW0, 1 s
   "SDC\DB_SDC_EMS_FLAGS\DB_SDC_EMS_FLAGS.EMS[139]" : Int AT %DB0.DBW0, 1 s
   "SDC\DB_SDC_EMS_FLAGS\DB_SDC_EMS_FLAGS.EMS[140]" : Int AT %DB0.DBW0, 1 s
   "SDC\DB_SDC_EMS_FLAGS\DB_SDC_EMS_FLAGS.EMS[141]" : Int AT %DB0.DBW0, 1 s
   "SDC\DB_SDC_EMS_FLAGS\DB_SDC_EMS_FLAGS.EMS[142]" : Int AT %DB0.DBW0, 1 s
   "SDC\DB_SDC_EMS_FLAGS\DB_SDC_EMS_FLAGS.EMS[143]" : Int AT %DB0.DBW0, 1 s
   "SDC\DB_SDC_EMS_FLAGS\DB_SDC_EMS_FLAGS.EMS[144]" : Int AT %DB0.DBW0, 1 s
   "SDC\DB_SDC_EMS_FLAGS\DB_SDC_EMS_FLAGS.EMS[145]" : Int AT %DB0.DBW0, 1 s
   "SDC\DB_SDC_EMS_FLAGS\DB_SDC_EMS_FLAGS.EMS[146]" : Int AT %DB0.DBW0, 1 s
   "SDC\DB_SDC_EMS_FLAGS\DB_SDC_EMS_FLAGS.EMS[147]" : Int AT %DB0.DBW0, 1 s
   "SDC\DB_SDC_EMS_FLAGS\DB_SDC_EMS_FLAGS.EMS[148]" : Int AT %DB0.DBW0, 1 s
   "SDC\DB_SDC_EMS_FLAGS\DB_SDC_EMS_FLAGS.EMS[149]" : Int AT %DB0.DBW0, 1 s
   "SDC\DB_SDC_EMS_FLAGS\DB_SDC_EMS_FLAGS.EMS[150]" : Int AT %DB0.DBW0, 1 s
   "SDC\DB_SDC_EMS_FLAGS\DB_SDC_EMS_FLAGS.EMS[151]" : Int AT %DB0.DBW0, 1 s
   "SDC\DB_SDC_EMS_FLAGS\DB_SDC_EMS_FLAGS.EMS[152]" : Int AT %DB0.DBW0, 1 s
   "SDC\DB_SDC_EMS_FLAGS\DB_SDC_EMS_FLAGS.EMS[153]" : Int AT %DB0.DBW0, 1 s
   "SDC\DB_SDC_EMS_FLAGS\DB_SDC_EMS_FLAGS.EMS[154]" : Int AT %DB0.DBW0, 1 s
   "SDC\DB_SDC_EMS_FLAGS\DB_SDC_EMS_FLAGS.EMS[155]" : Int AT %DB0.DBW0, 1 s
   "SDC\DB_SDC_EMS_FLAGS\DB_SDC_EMS_FLAGS.EMS[156]" : Int AT %DB0.DBW0, 1 s
   "SDC\DB_SDC_EMS_FLAGS\DB_SDC_EMS_FLAGS.EMS[157]" : Int AT %DB0.DBW0, 1 s
   "SDC\DB_SDC_EMS_FLAGS\DB_SDC_EMS_FLAGS.EMS[158]" : Int AT %DB0.DBW0, 1 s
   "SDC\DB_SDC_EMS_FLAGS\DB_SDC_EMS_FLAGS.EMS[159]" : Int AT %DB0.DBW0, 1 s
   "SDC\DB_SDC_EMS_FLAGS\DB_SDC_EMS_FLAGS.EMS[160]" : Int AT %DB0.DBW0, 1 s
   "SDC\DB_SDC_EMS_FLAGS\DB_SDC_EMS_FLAGS.EMS[161]" : Int AT %DB0.DBW0, 1 s
   "SDC\DB_SDC_EMS_FLAGS\DB_SDC_EMS_FLAGS.EMS[162]" : Int AT %DB0.DBW0, 1 s
   "SDC\DB_SDC_EMS_FLAGS\DB_SDC_EMS_FLAGS.EMS[163]" : Int AT %DB0.DBW0, 1 s
   "SDC\DB_SDC_EMS_FLAGS\DB_SDC_EMS_FLAGS.EMS[164]" : Int AT %DB0.DBW0, 1 s
   "SDC\DB_SDC_EMS_FLAGS\DB_SDC_EMS_FLAGS.EMS[165]" : Int AT %DB0.DBW0, 1 s
   "SDC\DB_SDC_EMS_FLAGS\DB_SDC_EMS_FLAGS.EMS[166]" : Int AT %DB0.DBW0, 1 s
   "SDC\DB_SDC_EMS_FLAGS\DB_SDC_EMS_FLAGS.EMS[167]" : Int AT %DB0.DBW0, 1 s
   "SDC\DB_SDC_EMS_FLAGS\DB_SDC_EMS_FLAGS.EMS[168]" : Int AT %DB0.DBW0, 1 s
   "SDC\DB_SDC_EMS_FLAGS\DB_SDC_EMS_FLAGS.EMS[169]" : Int AT %DB0.DBW0, 1 s
   "SDC\DB_SDC_EMS_FLAGS\DB_SDC_EMS_FLAGS.EMS[170]" : Int AT %DB0.DBW0, 1 s
   "SDC\DB_SDC_EMS_FLAGS\DB_SDC_EMS_FLAGS.EMS[171]" : Int AT %DB0.DBW0, 1 s
   "SDC\DB_SDC_EMS_FLAGS\DB_SDC_EMS_FLAGS.EMS[172]" : Int AT %DB0.DBW0, 1 s
   "SDC\DB_SDC_EMS_FLAGS\DB_SDC_EMS_FLAGS.EMS[173]" : Int AT %DB0.DBW0, 1 s
   "SDC\DB_SDC_EMS_FLAGS\DB_SDC_EMS_FLAGS.EMS[174]" : Int AT %DB0.DBW0, 1 s
   "SDC\DB_SDC_EMS_FLAGS\DB_SDC_EMS_FLAGS.EMS[175]" : Int AT %DB0.DBW0, 1 s
   "SDC\DB_SDC_EMS_FLAGS\DB_SDC_EMS_FLAGS.EMS[176]" : Int AT %DB0.DBW0, 1 s
   "SDC\DB_SDC_EMS_FLAGS\DB_SDC_EMS_FLAGS.EMS[177]" : Int AT %DB0.DBW0, 1 s
   "SDC\DB_SDC_EMS_FLAGS\DB_SDC_EMS_FLAGS.EMS[178]" : Int AT %DB0.DBW0, 1 s
   "SDC\DB_SDC_EMS_FLAGS\DB_SDC_EMS_FLAGS.EMS[179]" : Int AT %DB0.DBW0, 1 s
   "SDC\DB_SDC_EMS_FLAGS\DB_SDC_EMS_FLAGS.EMS[180]" : Int AT %DB0.DBW0, 1 s
   "SDC\DB_SDC_EMS_FLAGS\DB_SDC_EMS_FLAGS.EMS[181]" : Int AT %DB0.DBW0, 1 s
   "SDC\DB_SDC_EMS_FLAGS\DB_SDC_EMS_FLAGS.EMS[182]" : Int AT %DB0.DBW0, 1 s
   "SDC\DB_SDC_EMS_FLAGS\DB_SDC_EMS_FLAGS.EMS[183]" : Int AT %DB0.DBW0, 1 s
   "SDC\DB_SDC_EMS_FLAGS\DB_SDC_EMS_FLAGS.EMS[184]" : Int AT %DB0.DBW0, 1 s
